VERSION : 0.7
   VAR_INPUT
      MotorStarterID : Hw_Any;   // The ID of the motor starter to read the records from
      "FB Mode" : Int;
      ManualMode : Bool;   // Used only for FB_Mode = 1 / Manual Mode Signal
      AutoMode : Bool;   // Used only for FB_Mode = 1 / Auto Mode Signal
      Interlock : Bool;   // Interlock
      AutoOn : Bool;
      HandOn : Bool;   // Hand ON
      HandOff : Bool;   // Hand OFF
      SpareIN_1 : Bool;   // Spare
      RemoteFeedbackStat : Bool;   // Status - Remote Mode Feedback
      OnStatus : Bool;   // Status - On
      DeviceOStatus : Bool;   // Status - Device Ok
      CoolindDownPeriodStatus : Bool;   // Status - Cooling Down Period Active
      EmergencyStartExecStatus : Bool;   // Status - Emergency Start Executed
      GeneralWarningStatus : Bool;   // Fault - General Warning
      GeneralFaultStatus : Bool;   // Fault - General Fault
      OverloadOperationEvent : Bool;   // Event - Overload Operation Fault (I>115%Is)
      OverloadFaultEvent : Bool;   // Event - Overload Fault
      UnbalanceFault : Bool;   // Event - Unbalance Fault
      OLandLossOfPhaseEvent : Bool;   // Event - Overload and Loss of Phase
      StalledRotorEvent : Bool;   // Event - Stalled Rotor
      HardwareFaultBasicUnitTrip : Bool;   // Trip - Hardware Fault Basic Unit
      ModuleFaultTrip : Bool;   // Trip - Module Fault
      ExecOnCommandTrip : Bool;   // Trip - Execution On-Command
      RemainingCooldDownPeriod : Int;   // Remaining Cool Down Period
      FullLoadAmps : Real;   // Full Load Amps
   END_VAR
   VAR_OUTPUT
      SpareOUT_1 : Bool;
      Stop_CMD : Bool;   // Stop Command for the Semicode
      Start_CMD : Bool;   // Start Command for the Semicode
      TestSimocode : Bool;   // Simocode Test
      EmergenyStart : Bool;   // Emergency Start
      RemoteCommandsEnabled : Bool;   // Auto Mode / Enable Remote Commands
      ResetSimocode : Bool;   // Simocode Reset
      SpareOUT_2 : Bool;
      SpareOUT_3 : Bool;
      SpareOUT_4 : Bool;
      SpareOUT_5 : Bool;
      SpareOUT_6 : Bool;
      SpareOUT_7 : Bool;
      SpareOUT_8 : Bool;
      SpareOUT_9 : Bool;
      SpareOUT_10 : Bool;
      SpareOUTW_1 : Int;
      SpareOUTW_2 : Int;
   END_VAR
   VAR
      HMI : Struct
         Controls : Struct
            Start : Bool;
            Stop : Bool;
            Reset : Bool;
            PLCMOHR : Bool;   // PLC Motor Operating Hours Reset
         END_STRUCT;
         Status : Struct
            Mode : Int;   // Simocode Mode
            MotorOperatingHours : Real;   // True Semicode Motor Operating Hours
            DeviceOperatingHours : Real;
            LMOH : Real;   // Last Motor Operating Hours
            RemainingCoolDownPeriod : Int;   // Remaining Cooldown Period
            MaxNumberOLtrips : Int;   // Maximum Number of Overload Trips
            ControlStatusWord : Word;   // Control/Status Information Bits
            MaxCurrent : Real;   // Maximum Current (Is %)
            Current1 : Real;   // Leg 1 Current (Is %)
            Current2 : Real;   // Leg 2 Current (Is %)
            Current3 : Real;   // Leg 3 Current (Is %)
            LastTripCurrent : Real;   // Last Trip Current (% of Is)
            CommandSimocode : Bool;   // Commanding Simocode to Start
         END_STRUCT;
         Config : Struct
            "RemainingCoolDownPeriod.SP" : Int := 300;
            Start_PT : Time := T#500MS;
            Stop_PT : Time := T#500MS;
         END_STRUCT;
         Math : Struct
            MOH1 : DInt;
            MOH2 : Real;
            PLCMOH : Real;   // PLC Motor Operating Hours
            LMOH : Real;
         END_STRUCT;
      END_STRUCT;
      OS : Struct
         RON : Bool;   // Remote / HMI On
         ROFF : Bool;   // Remote / HMI Off
         HON : Bool;   // Hand/Local On
         HOFF : Bool;   // Hand/Local Off
         PLCMOHR : Bool;
         LMOH1 : Bool;
         LMOH2 : Bool;
         RST : Bool;   // Reset Semicode
      END_STRUCT;
      "DS94 Record" : Struct
         "Phase Current L1 %" : USInt;
         "Phase Current L2 %" : USInt;
         "Phase Current L3 %" : USInt;
         Reserved_3 : Byte;
         "Remaining cool-down time of the motor" : UInt;
         "Motor heating_6" : USInt;
         Unbalance : USInt;
         "Motor Heating" : UInt;
         Reserved_10 : Byte;
         Reserved_11 : Byte;
         Reserved_12 : Byte;
         Reserved_13 : Byte;
         Reserved_14 : Byte;
         Reserved_15 : Byte;
         Reserved_16 : Byte;
         Reserved_17 : Byte;
         Reserved_18 : Byte;
         Reserved_19 : Byte;
         Reserved_20 : Byte;
         Reserved_21 : Byte;
         Reserved_22 : Byte;
         Reserved_23 : Byte;
         Reserved_24 : Byte;
         Reserved_25 : Byte;
         Reserved_26 : Byte;
         Reserved_27 : Byte;
         "Phase Current L1 (rms)" : UDInt;
         "Phase Current L2 (rms)" : UDInt;
         "Phase Current L3 (rms)" : UDInt;
         "Electronics Supply Voltage" : UInt;
         Reserved_42 : Byte;
         Reserved_43 : Byte;
         Reserved_44 : Byte;
         Reserved_45 : Byte;
         Reserved_46 : Byte;
         Reserved_47 : Byte;
         Reserved_48 : Byte;
         Reserved_49 : Byte;
         Reserved_50 : Byte;
         Reserved_51 : Byte;
         Reserved_52 : Byte;
         Reserved_53 : Byte;
         Reserved_54 : Byte;
         Reserved_55 : Byte;
         Reserved_56 : Byte;
         Reserved_57 : Byte;
         Reserved_58 : Byte;
         Reserved_59 : Byte;
         Reserved_60 : Byte;
         Reserved_61 : Byte;
         Reserved_62 : Byte;
         Reserved_63 : Byte;
      END_STRUCT;
      "DS94 Record_1" : Struct
         "Phase Current L1 %" : USInt;
         "Phase Current L2 %" : USInt;
         "Phase Current L3 %" : USInt;
         Reserved_3 : Byte;
         "Remaining cool-down time of the motor" : UInt;
         "Motor heating_6" : USInt;
         "Asymmetry value_7" : USInt;
         Reserved_8 : Byte;
         Reserved_9 : Byte;
         Reserved_10 : Byte;
         Reserved_11 : Byte;
         Reserved_12 : Byte;
         Reserved_13 : Byte;
         Reserved_14 : Byte;
         Reserved_15 : Byte;
         Reserved_16 : Byte;
         Reserved_17 : Byte;
         Reserved_18 : Byte;
         Reserved_19 : Byte;
         Reserved_20 : Byte;
         Reserved_21 : Byte;
         Reserved_22 : Byte;
         Reserved_23 : Byte;
         Reserved_24 : Byte;
         Reserved_25 : Byte;
         Reserved_26 : Byte;
         Reserved_27 : Byte;
         "Phase Current L1 (rms)" : UDInt;
         "Phase Current L2 (rms)" : UDInt;
         "Phase Current L3 (rms)" : UDInt;
         "Electronics Supply Voltage" : USInt;
         Reserved_46 : Byte;
         Reserved_47 : Byte;
         Reserved_48 : Byte;
         Reserved_49 : Byte;
         Reserved_50 : Byte;
         Reserved_51 : Byte;
         Reserved_52 : Byte;
         Reserved_53 : Byte;
         Reserved_54 : Byte;
         Reserved_55 : Byte;
         Reserved_56 : Byte;
         Reserved_57 : Byte;
         Reserved_58 : Byte;
         Reserved_59 : Byte;
         Reserved_60 : Byte;
         Reserved_61 : Byte;
         Reserved_62 : Byte;
      END_STRUCT;
      "DS95 Record" : Struct
         Reserved_0 : USInt;
         "Reserved_1.0" : Bool;
         "Reserved_1.1" : Bool;
         "Reserved_1.2" : Bool;
         "Reserved_1.3" : Bool;
         "Reserved_1.4" : Bool;
         "Reserved_1.5" : Bool;
         "Reserved_1.6" : Bool;
         "Reserved_1.7" : Bool;
         Reserved_2 : Byte;
         Reserved_3 : Byte;
         "Device operating hours in seconds" : UDInt;
         "Number of motor CW starts" : UDInt;
         "Number of starts motor CCW" : UDInt;
         "Number of motor overload trips" : UInt;
         Reserved_18 : Byte;
         Reserved_19 : Byte;
         "Motor current_20..23" : UDInt;
         "Last tripping current_24..27" : DInt;
         "Motor operating hours in seconds_28...31" : UDInt;
         Reserved_32 : Byte;
         Reserved_33 : Byte;
         Reserved_34 : Byte;
         Reserved_35 : Byte;
         Reserved_36 : Byte;
         Reserved_37 : Byte;
         Reserved_38 : Byte;
         Reserved_39 : Byte;
         Reserved_40 : Byte;
         Reserved_41 : Byte;
         Reserved_42 : Byte;
         Reserved_43 : Byte;
         Reserved_44 : Byte;
         Reserved_45 : Byte;
         Reserved_46 : Byte;
         Reserved_47 : Byte;
         Reserved_48 : Byte;
         Reserved_49 : Byte;
         "Number of switching element" : UInt;
         "Number of hard switching" : UInt;
         Reserved_54 : Byte;
         Reserved_55 : Byte;
         Reserved_56 : Byte;
         Reserved_57 : Byte;
         Reserved_58 : Byte;
         Reserved_59 : Byte;
         Reserved_60 : Byte;
         Reserved_61 : Byte;
         Reserved_62 : Byte;
         Reserved_63 : Byte;
         Reserved_64 : Byte;
         Reserved_65 : Byte;
         Reserved_66 : Byte;
         Reserved_67 : Byte;
         Reserved_68 : Byte;
         Reserved_69 : Byte;
         Reserved_70 : Byte;
         Reserved_71 : Byte;
         Reserved_72 : Byte;
         Reserved_73 : Byte;
         Reserved_74 : Byte;
         Reserved_75 : Byte;
         Reserved_76 : Byte;
         Reserved_77 : Byte;
         Reserved_78 : Byte;
         Reserved_79 : Byte;
         Reserved_80 : Byte;
         Reserved_81 : Byte;
         Reserved_82 : Byte;
         Reserved_83 : Byte;
         Reserved_84 : Byte;
         Reserved_85 : Byte;
         Reserved_86 : Byte;
         Reserved_87 : Byte;
         Reserved_88 : Byte;
         Reserved_89 : Byte;
      END_STRUCT;
      START_CMD_TOF : TOF_TIME;   // Start Semicode
      STOP_CMD_TOF : TOF_TIME;
      Current_RDREC : RDREC;
      Time_RDREC : RDREC;
      RDREC_REQ : SInt;
      Current_Error : SInt;
      Time_Error : SInt;
      flnk : Array[0..2] of Bool;
   END_VAR
   VAR_TEMP
      IL1_Math2 : Real;
      IL1_Math3 : Real;
      IL2_Math2 : Real;
      IL2_Math3 : Real;
      IL3_Math2 : Real;
      IL3_Math3 : Real;
      MC_Math1 : DInt;
      MC_Math2 : Real;
      MC_Math3 : Real;
      LTC_Math2 : Real;
      LTC_Math3 : Real;
      Start : Bool;
      Fault : Bool;
      "Valid Current" : Bool;
      "Valid Time" : Bool;
      MOTS : Real;   // Motor Operating Time in Seconds
      DOTH : Real;   // Device Operating Time in Hours
      DOTS : Real;   // Device Operating Time in Seconds
      MOTH : Real;   // Motor Operating Time in hours
   END_VAR
   VAR_TEMP   // added for the SCL form of the ladder/FBD networks
      _w1 : Bool;
      _w2 : Bool;
      _w3 : Bool;
      _w4 : Bool;
      _w5 : Bool;
   END_VAR
BEGIN

REGION Network 1: Read request
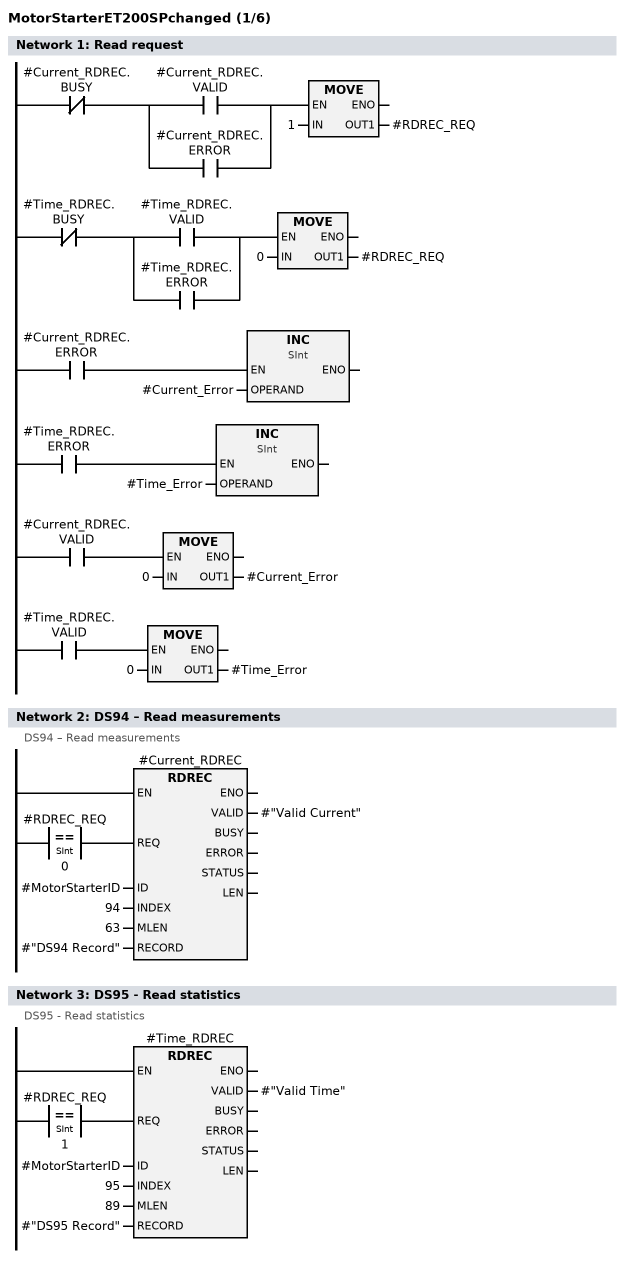
   RUNG wire#powerrail
      I_Contact( #Current_RDREC.BUSY )
      wire#w1
      Contact( #Current_RDREC.VALID )
      wire#w2
      Move(in := 1, out1 => #RDREC_REQ)
   END_RUNG
   RUNG wire#w1
      Contact( #Current_RDREC.ERROR )
   END_RUNG wire#w2
   RUNG wire#powerrail
      I_Contact( #Time_RDREC.BUSY )
      wire#w3
      Contact( #Time_RDREC.VALID )
      wire#w4
      Move(in := 0, out1 => #RDREC_REQ)
   END_RUNG
   RUNG wire#w3
      Contact( #Time_RDREC.ERROR )
   END_RUNG wire#w4
   RUNG wire#powerrail
      Contact( #Current_RDREC.ERROR )
      { S7_Templates := "DestType := SInt" } Inc( #Current_Error )
   END_RUNG
   RUNG wire#powerrail
      Contact( #Time_RDREC.ERROR )
      { S7_Templates := "DestType := SInt" } Inc( #Time_Error )
   END_RUNG
   RUNG wire#powerrail
      Contact( #Current_RDREC.VALID )
      Move(in := 0, out1 => #Current_Error)
   END_RUNG
   RUNG wire#powerrail
      Contact( #Time_RDREC.VALID )
      Move(in := 0, out1 => #Time_Error)
   END_RUNG
   // the same network as SCL:
   IF NOT #Current_RDREC.BUSY AND (#Current_RDREC.VALID OR #Current_RDREC.ERROR) THEN
       #RDREC_REQ := 1;
   END_IF;
   IF NOT #Time_RDREC.BUSY AND (#Time_RDREC.VALID OR #Time_RDREC.ERROR) THEN #RDREC_REQ := 0; END_IF;
   IF #Current_RDREC.ERROR THEN #Current_Error := #Current_Error + 1; END_IF;
   IF #Time_RDREC.ERROR THEN #Time_Error := #Time_Error + 1; END_IF;
   IF #Current_RDREC.VALID THEN #Current_Error := 0; END_IF;
   IF #Time_RDREC.VALID THEN #Time_Error := 0; END_IF;
END_REGION

REGION Network 2: DS94 – Read measurements
   // DS94 – Read measurements
   #Current_RDREC(REQ := #RDREC_REQ = 0,   // RDREC
                  ID := #MotorStarterID,
                  INDEX := 94,
                  MLEN := 63,
                  RECORD := #"DS94 Record",
                  VALID => #"Valid Current");
END_REGION

REGION Network 3: DS95 - Read statistics
   // DS95 - Read statistics
   #Time_RDREC(REQ := #RDREC_REQ = 1,   // RDREC
               ID := #MotorStarterID,
               INDEX := 95,
               MLEN := 89,
               RECORD := #"DS95 Record",
               VALID => #"Valid Time");
END_REGION

REGION Network 4: HOA in Off
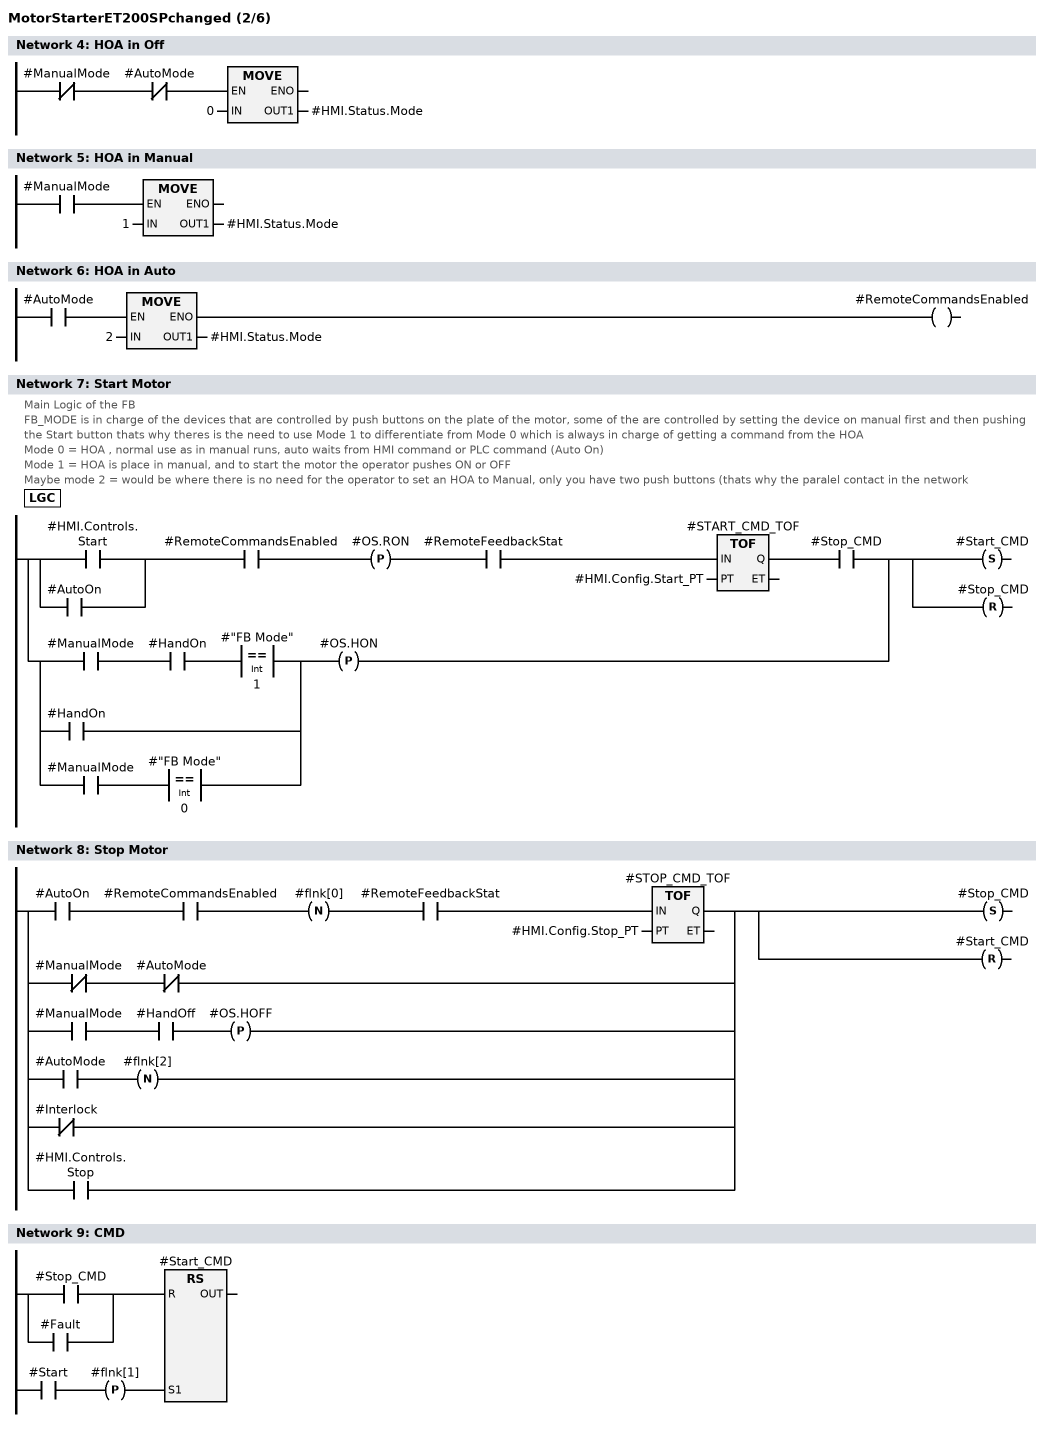
   RUNG wire#powerrail
      I_Contact( #ManualMode )
      I_Contact( #AutoMode )
      { S7_GenerateENO := "TRUE" } Move(in := 0, out1 => #HMI.Status.Mode)
   END_RUNG
   // the same network as SCL:
   IF NOT #ManualMode AND NOT #AutoMode THEN #HMI.Status.Mode := 0; END_IF;
END_REGION

REGION Network 5: HOA in Manual
   RUNG wire#powerrail
      Contact( #ManualMode )
      { S7_GenerateENO := "TRUE" } Move(in := 1, out1 => #HMI.Status.Mode)
   END_RUNG
   // the same network as SCL:
   IF #ManualMode THEN #HMI.Status.Mode := 1; END_IF;
END_REGION

REGION Network 6: HOA in Auto
   RUNG wire#powerrail
      Contact( #AutoMode )
      { S7_GenerateENO := "TRUE" } Move(in := 2, out1 => #HMI.Status.Mode)
      Coil( #RemoteCommandsEnabled )
   END_RUNG
   // the same network as SCL:
   // ENO of a box is taken as its EN; it also drops when the box reports an error
   IF #AutoMode THEN #HMI.Status.Mode := 2; END_IF;
   #RemoteCommandsEnabled := #AutoMode;
END_REGION

REGION Network 7: Start Motor
   // Main Logic of the FB
   // FB_MODE is in charge of the devices that are controlled by push buttons on the plate of the motor, some of the are controlled by setting the device on manual first and then pushing the Start button thats why theres is the need to use Mode 1 to differentiate from Mode 0 which is always in charge of getting a command from the HOA
   // Mode 0 = HOA , normal use as in manual runs, auto waits from HMI command or PLC command (Auto On)
   // Mode 1 = HOA is place in manual, and to start the motor the operator pushes ON or OFF
   // Maybe mode 2 = would be where there is no need for the operator to set an HOA to Manual, only you have two push buttons (thats why the paralel contact in the network
   LGC:
   #_w1 := (#HMI.Controls.Start OR #AutoOn) AND #RemoteCommandsEnabled;
   #_w2 := #_w1 AND NOT #OS.RON;   // rising edge
   #OS.RON := #_w1;
   #START_CMD_TOF(IN := #_w2 AND #RemoteFeedbackStat, PT := #HMI.Config.Start_PT);   // TOF
   #_w3 := (#ManualMode AND #HandOn AND (#"FB Mode" = 1)) OR #HandOn OR (#ManualMode AND (#"FB Mode" = 0));
   #_w4 := #_w3 AND NOT #OS.HON;   // rising edge
   #OS.HON := #_w3;
   IF (#START_CMD_TOF.Q AND #Stop_CMD) OR #_w4 THEN
       #Start_CMD := TRUE;
       #Stop_CMD := FALSE;
   END_IF;
END_REGION

REGION Network 8: Stop Motor
   #_w1 := #AutoOn AND #RemoteCommandsEnabled;
   #_w2 := NOT #_w1 AND #flnk[0];   // falling edge
   #flnk[0] := #_w1;
   #STOP_CMD_TOF(IN := #_w2 AND #RemoteFeedbackStat, PT := #HMI.Config.Stop_PT);   // TOF
   #_w3 := #ManualMode AND #HandOff;
   #_w4 := #_w3 AND NOT #OS.HOFF;   // rising edge
   #OS.HOFF := #_w3;
   #_w5 := NOT #AutoMode AND #flnk[2];   // falling edge
   #flnk[2] := #AutoMode;
   IF #STOP_CMD_TOF.Q OR (NOT #ManualMode AND NOT #AutoMode) OR #_w4 OR #_w5 OR NOT #Interlock OR #HMI.Controls.Stop THEN
       #Stop_CMD := TRUE;
       #Start_CMD := FALSE;
   END_IF;
END_REGION

REGION Network 9: CMD
   RUNG wire#powerrail
      Contact( #Stop_CMD )
      wire#w1
      S_RS(operand := #Start_CMD, s1 := wire#w2)
   END_RUNG
   RUNG wire#powerrail
      Contact( #Fault )
   END_RUNG wire#w1
   RUNG wire#powerrail
      Contact( #Start )
      P_Trig( #flnk[1] )
   END_RUNG wire#w2
   // the same network as SCL:
   #_w1 := #Start AND NOT #flnk[1];   // rising edge
   #flnk[1] := #Start;
   IF #Stop_CMD OR #Fault THEN
       #Start_CMD := FALSE;   // RS flip-flop
   END_IF;
   IF #_w1 THEN #Start_CMD := TRUE; END_IF;
END_REGION

REGION Network 10: Interlock
   // Main Logic of the FB
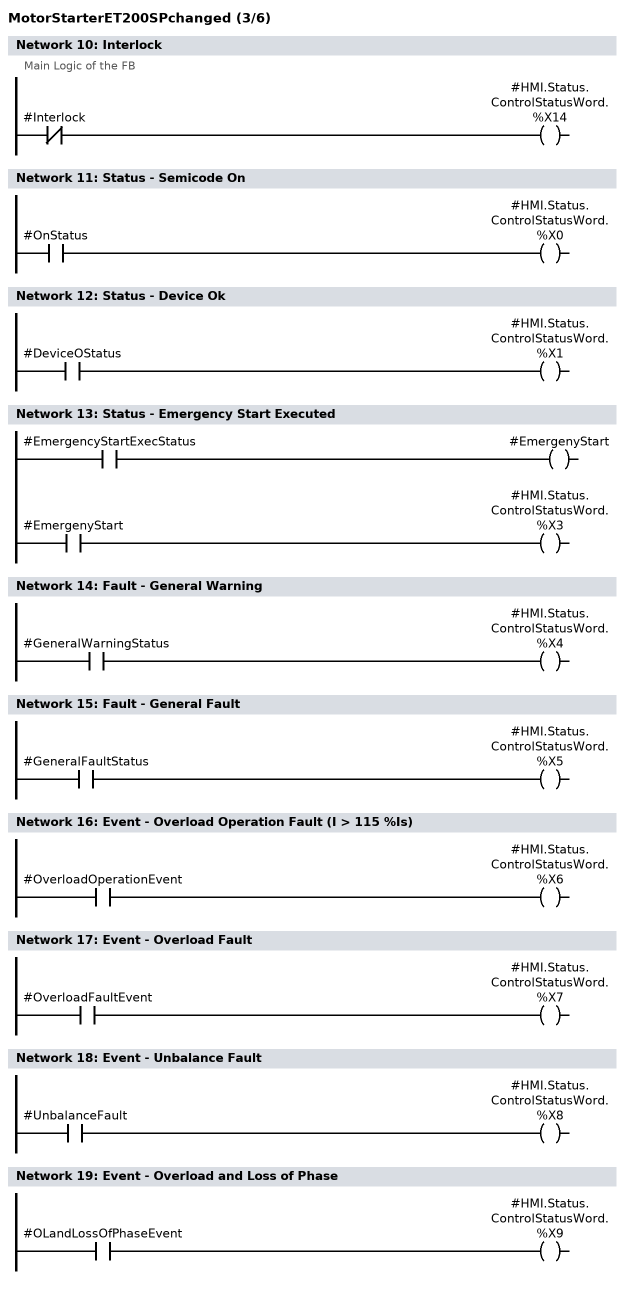
   RUNG wire#powerrail
      I_Contact( #Interlock )
      Coil( #HMI.Status.ControlStatusWord.%X14 )
   END_RUNG
   // the same network as SCL:
   #HMI.Status.ControlStatusWord.%X14 := NOT #Interlock;
END_REGION

REGION Network 11: Status - Semicode On
   RUNG wire#powerrail
      Contact( #OnStatus )
      Coil( #HMI.Status.ControlStatusWord.%X0 )
   END_RUNG
   // the same network as SCL:
   #HMI.Status.ControlStatusWord.%X0 := #OnStatus;
END_REGION

REGION Network 12: Status - Device Ok
   RUNG wire#powerrail
      Contact( #DeviceOStatus )
      Coil( #HMI.Status.ControlStatusWord.%X1 )
   END_RUNG
   // the same network as SCL:
   #HMI.Status.ControlStatusWord.%X1 := #DeviceOStatus;
END_REGION

REGION Network 13: Status - Emergency Start Executed
   RUNG wire#powerrail
      Contact( #EmergencyStartExecStatus )
      Coil( #EmergenyStart )
   END_RUNG
   RUNG wire#powerrail
      Contact( #EmergenyStart )
      Coil( #HMI.Status.ControlStatusWord.%X3 )
   END_RUNG
   // the same network as SCL:
   #EmergenyStart := #EmergencyStartExecStatus;
   #HMI.Status.ControlStatusWord.%X3 := #EmergenyStart;
END_REGION

REGION Network 14: Fault - General Warning
   RUNG wire#powerrail
      Contact( #GeneralWarningStatus )
      Coil( #HMI.Status.ControlStatusWord.%X4 )
   END_RUNG
   // the same network as SCL:
   #HMI.Status.ControlStatusWord.%X4 := #GeneralWarningStatus;
END_REGION

REGION Network 15: Fault - General Fault
   RUNG wire#powerrail
      Contact( #GeneralFaultStatus )
      Coil( #HMI.Status.ControlStatusWord.%X5 )
   END_RUNG
   // the same network as SCL:
   #HMI.Status.ControlStatusWord.%X5 := #GeneralFaultStatus;
END_REGION

REGION Network 16: Event - Overload Operation Fault (I > 115 %Is)
   RUNG wire#powerrail
      Contact( #OverloadOperationEvent )
      Coil( #HMI.Status.ControlStatusWord.%X6 )
   END_RUNG
   // the same network as SCL:
   #HMI.Status.ControlStatusWord.%X6 := #OverloadOperationEvent;
END_REGION

REGION Network 17: Event - Overload Fault
   RUNG wire#powerrail
      Contact( #OverloadFaultEvent )
      Coil( #HMI.Status.ControlStatusWord.%X7 )
   END_RUNG
   // the same network as SCL:
   #HMI.Status.ControlStatusWord.%X7 := #OverloadFaultEvent;
END_REGION

REGION Network 18: Event - Unbalance Fault
   RUNG wire#powerrail
      Contact( #UnbalanceFault )
      Coil( #HMI.Status.ControlStatusWord.%X8 )
   END_RUNG
   // the same network as SCL:
   #HMI.Status.ControlStatusWord.%X8 := #UnbalanceFault;
END_REGION

REGION Network 19: Event - Overload and Loss of Phase
   RUNG wire#powerrail
      Contact( #OLandLossOfPhaseEvent )
      Coil( #HMI.Status.ControlStatusWord.%X9 )
   END_RUNG
   // the same network as SCL:
   #HMI.Status.ControlStatusWord.%X9 := #OLandLossOfPhaseEvent;
END_REGION

REGION Network 20: Event - Stalled Rotor
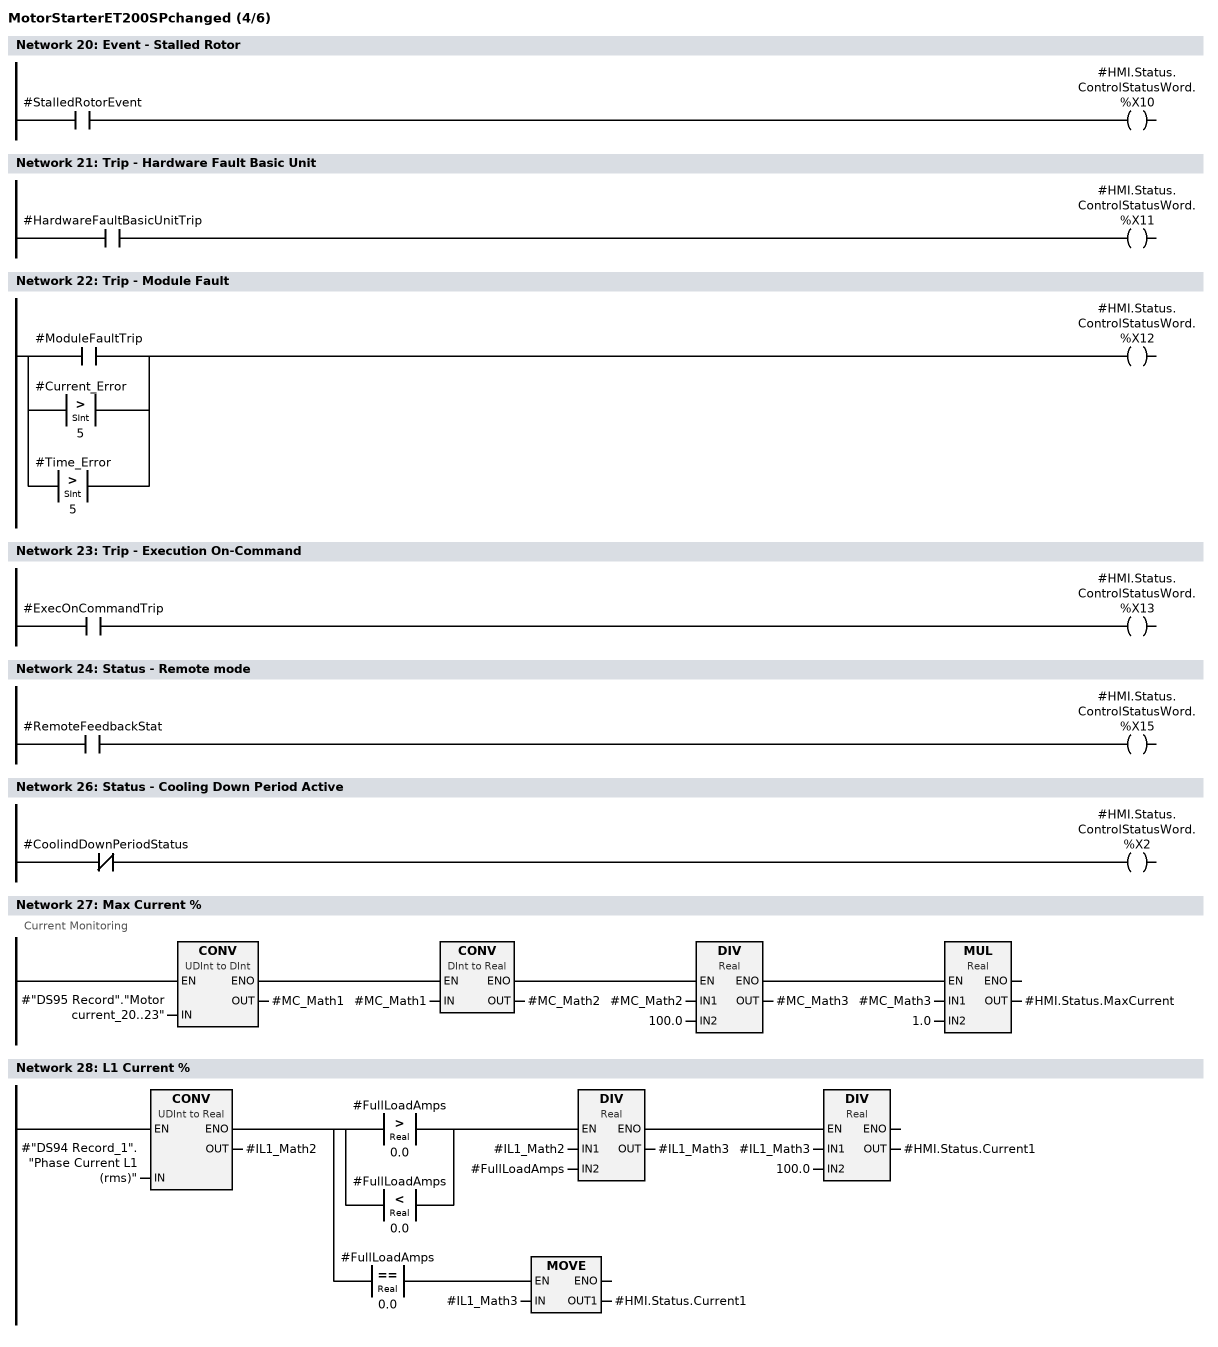
   RUNG wire#powerrail
      Contact( #StalledRotorEvent )
      Coil( #HMI.Status.ControlStatusWord.%X10 )
   END_RUNG
   // the same network as SCL:
   #HMI.Status.ControlStatusWord.%X10 := #StalledRotorEvent;
END_REGION

REGION Network 21: Trip - Hardware Fault Basic Unit
   RUNG wire#powerrail
      Contact( #HardwareFaultBasicUnitTrip )
      Coil( #HMI.Status.ControlStatusWord.%X11 )
   END_RUNG
   // the same network as SCL:
   #HMI.Status.ControlStatusWord.%X11 := #HardwareFaultBasicUnitTrip;
END_REGION

REGION Network 22: Trip - Module Fault
   RUNG wire#powerrail
      Contact( #ModuleFaultTrip )
      wire#w1
      Coil( #HMI.Status.ControlStatusWord.%X12 )
   END_RUNG
   RUNG wire#powerrail
      { S7_Templates := "SrcType := SInt" } GT_Contact(in1 := #Current_Error, in2 := 5)
   END_RUNG wire#w1
   RUNG wire#powerrail
      { S7_Templates := "SrcType := SInt" } GT_Contact(in1 := #Time_Error, in2 := 5)
   END_RUNG wire#w1
   // the same network as SCL:
   #HMI.Status.ControlStatusWord.%X12 := #ModuleFaultTrip OR (#Current_Error > 5) OR (#Time_Error > 5);
END_REGION

REGION Network 23: Trip - Execution On-Command
   RUNG wire#powerrail
      Contact( #ExecOnCommandTrip )
      Coil( #HMI.Status.ControlStatusWord.%X13 )
   END_RUNG
   // the same network as SCL:
   #HMI.Status.ControlStatusWord.%X13 := #ExecOnCommandTrip;
END_REGION

REGION Network 24: Status - Remote mode
   RUNG wire#powerrail
      Contact( #RemoteFeedbackStat )
      Coil( #HMI.Status.ControlStatusWord.%X15 )
   END_RUNG
   // the same network as SCL:
   #HMI.Status.ControlStatusWord.%X15 := #RemoteFeedbackStat;
END_REGION

REGION Network 25 (SCL): Motor Operating Hours
   #DOTS := UDINT_TO_REAL(#"DS95 Record"."Device operating hours in seconds");
   #DOTH := #DOTS / Real#3610.68;
   #MOTS := UDINT_TO_REAL(#"DS95 Record"."Motor operating hours in seconds_28...31");
   #MOTH := #MOTS / Real#6027.66;
   #HMI.Status.DeviceOperatingHours := #DOTH;
   #HMI.Status.MotorOperatingHours := #MOTH;
END_REGION

REGION Network 26: Status - Cooling Down Period Active
   RUNG wire#powerrail
      I_Contact( #CoolindDownPeriodStatus )
      Coil( #HMI.Status.ControlStatusWord.%X2 )
   END_RUNG
   // the same network as SCL:
   #HMI.Status.ControlStatusWord.%X2 := NOT #CoolindDownPeriodStatus;
END_REGION

REGION Network 27: Max Current %
   // Current Monitoring
   RUNG wire#powerrail
      { S7_Templates := "[SrcType := UDInt, DestType := DInt]"; S7_GenerateENO := "TRUE" } Convert(in := #"DS95 Record"."Motor current_20..23", out => #MC_Math1)
      { S7_Templates := "[SrcType := DInt, DestType := Real]"; S7_GenerateENO := "TRUE" } Convert(in := #MC_Math1, out => #MC_Math2)
      { S7_Templates := "SrcType := Real"; S7_GenerateENO := "TRUE" } Div(in1 := #MC_Math2, in2 := 100.0, out => #MC_Math3)
      { S7_Templates := "SrcType := Real"; S7_GenerateENO := "TRUE" } Mul(in1 := #MC_Math3, in2 := 1.0, out => #HMI.Status.MaxCurrent)
   END_RUNG
   // the same network as SCL:
   // ENO of a box is taken as its EN; it also drops when the box reports an error
   #MC_Math1 := UDINT_TO_DINT(#"DS95 Record"."Motor current_20..23");
   #MC_Math2 := DINT_TO_REAL(#MC_Math1);
   #MC_Math3 := #MC_Math2 / 100.0;
   #HMI.Status.MaxCurrent := #MC_Math3 * 1.0;
END_REGION

REGION Network 28: L1 Current %
   RUNG wire#powerrail
      { S7_Templates := "[SrcType := UDInt, DestType := Real]"; S7_GenerateENO := "TRUE" } Convert(in := #"DS94 Record_1"."Phase Current L1 (rms)", out => #IL1_Math2)
      wire#w1
      { S7_Templates := "SrcType := Real" } GT_Contact(in1 := #FullLoadAmps, in2 := 0.0)
      wire#w2
      { S7_Templates := "SrcType := Real"; S7_GenerateENO := "TRUE" } Div(in1 := #IL1_Math2, in2 := #FullLoadAmps, out => #IL1_Math3)
      { S7_Templates := "SrcType := Real"; S7_GenerateENO := "TRUE" } Div(in1 := #IL1_Math3, in2 := 100.0, out => #HMI.Status.Current1)
   END_RUNG
   RUNG wire#w1
      { S7_Templates := "SrcType := Real" } LT_Contact(in1 := #FullLoadAmps, in2 := 0.0)
   END_RUNG wire#w2
   RUNG wire#w1
      { S7_Templates := "SrcType := Real" } EQ_Contact(in1 := #FullLoadAmps, in2 := 0.0)
      Move(in := #IL1_Math3, out1 => #HMI.Status.Current1)
   END_RUNG
   // the same network as SCL:
   // ENO of a box is taken as its EN; it also drops when the box reports an error
   #IL1_Math2 := UDINT_TO_REAL(#"DS94 Record_1"."Phase Current L1 (rms)");
   IF (#FullLoadAmps > 0.0) OR (#FullLoadAmps < 0.0) THEN
       #IL1_Math3 := #IL1_Math2 / #FullLoadAmps;
       #HMI.Status.Current1 := #IL1_Math3 / 100.0;
   END_IF;
   IF #FullLoadAmps = 0.0 THEN #HMI.Status.Current1 := #IL1_Math3; END_IF;
END_REGION

REGION Network 29: L2 Current %
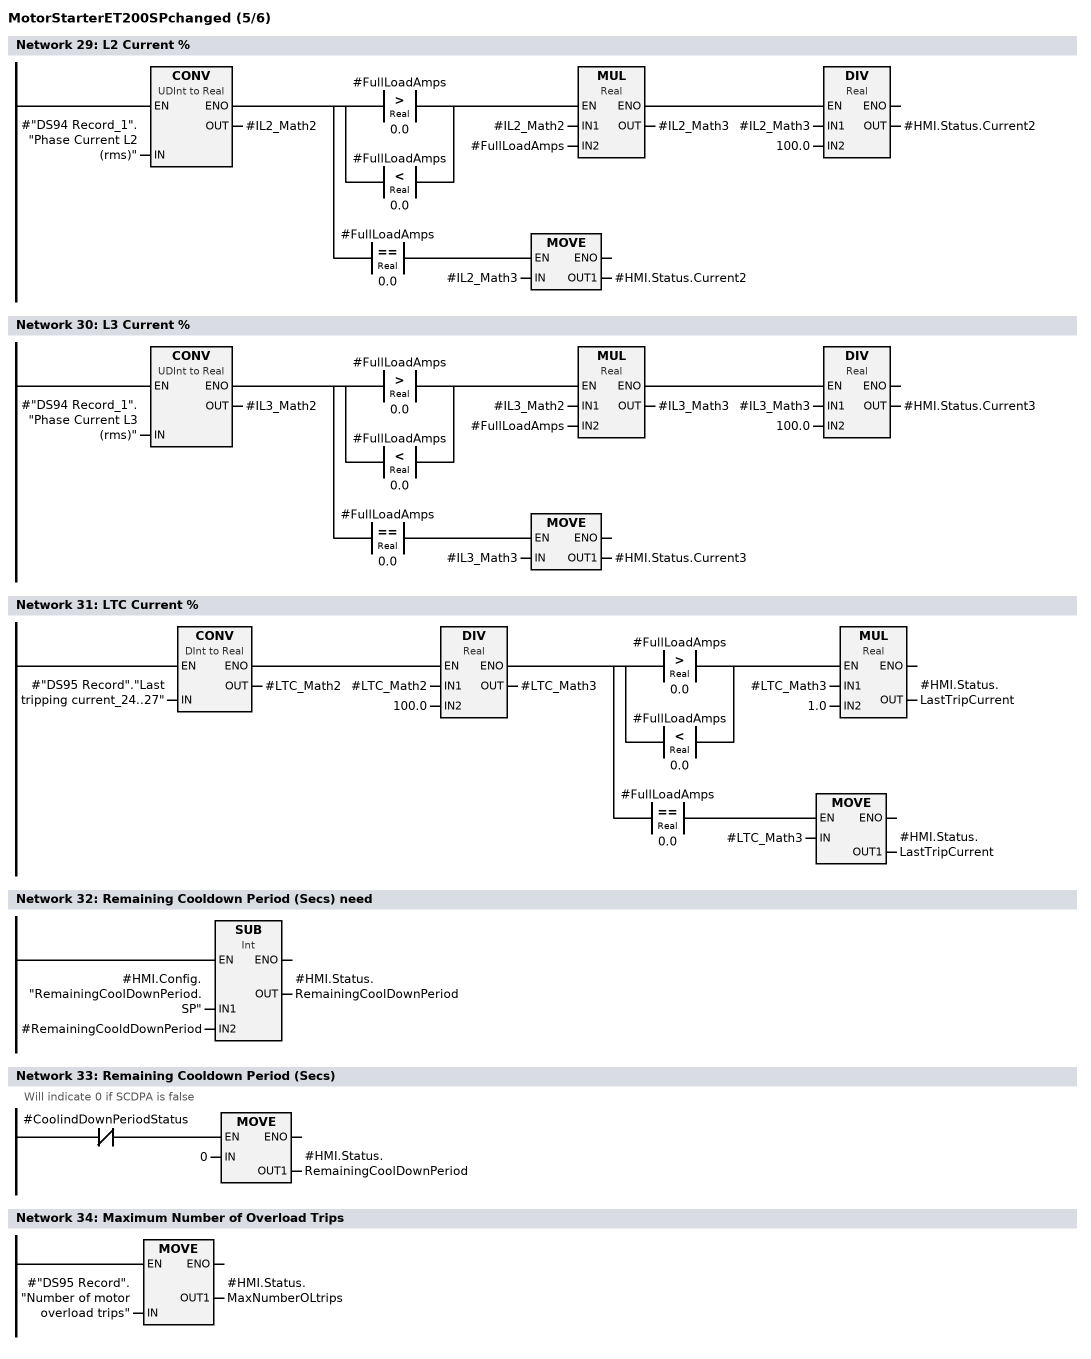
   RUNG wire#powerrail
      { S7_Templates := "[SrcType := UDInt, DestType := Real]"; S7_GenerateENO := "TRUE" } Convert(in := #"DS94 Record_1"."Phase Current L2 (rms)", out => #IL2_Math2)
      wire#w1
      { S7_Templates := "SrcType := Real" } GT_Contact(in1 := #FullLoadAmps, in2 := 0.0)
      wire#w2
      { S7_Templates := "SrcType := Real"; S7_GenerateENO := "TRUE" } Mul(in1 := #IL2_Math2, in2 := #FullLoadAmps, out => #IL2_Math3)
      { S7_Templates := "SrcType := Real"; S7_GenerateENO := "TRUE" } Div(in1 := #IL2_Math3, in2 := 100.0, out => #HMI.Status.Current2)
   END_RUNG
   RUNG wire#w1
      { S7_Templates := "SrcType := Real" } LT_Contact(in1 := #FullLoadAmps, in2 := 0.0)
   END_RUNG wire#w2
   RUNG wire#w1
      { S7_Templates := "SrcType := Real" } EQ_Contact(in1 := #FullLoadAmps, in2 := 0.0)
      Move(in := #IL2_Math3, out1 => #HMI.Status.Current2)
   END_RUNG
   // the same network as SCL:
   // ENO of a box is taken as its EN; it also drops when the box reports an error
   #IL2_Math2 := UDINT_TO_REAL(#"DS94 Record_1"."Phase Current L2 (rms)");
   IF (#FullLoadAmps > 0.0) OR (#FullLoadAmps < 0.0) THEN
       #IL2_Math3 := #IL2_Math2 * #FullLoadAmps;
       #HMI.Status.Current2 := #IL2_Math3 / 100.0;
   END_IF;
   IF #FullLoadAmps = 0.0 THEN #HMI.Status.Current2 := #IL2_Math3; END_IF;
END_REGION

REGION Network 30: L3 Current %
   RUNG wire#powerrail
      { S7_Templates := "[SrcType := UDInt, DestType := Real]"; S7_GenerateENO := "TRUE" } Convert(in := #"DS94 Record_1"."Phase Current L3 (rms)", out => #IL3_Math2)
      wire#w1
      { S7_Templates := "SrcType := Real" } GT_Contact(in1 := #FullLoadAmps, in2 := 0.0)
      wire#w2
      { S7_Templates := "SrcType := Real"; S7_GenerateENO := "TRUE" } Mul(in1 := #IL3_Math2, in2 := #FullLoadAmps, out => #IL3_Math3)
      { S7_Templates := "SrcType := Real"; S7_GenerateENO := "TRUE" } Div(in1 := #IL3_Math3, in2 := 100.0, out => #HMI.Status.Current3)
   END_RUNG
   RUNG wire#w1
      { S7_Templates := "SrcType := Real" } LT_Contact(in1 := #FullLoadAmps, in2 := 0.0)
   END_RUNG wire#w2
   RUNG wire#w1
      { S7_Templates := "SrcType := Real" } EQ_Contact(in1 := #FullLoadAmps, in2 := 0.0)
      Move(in := #IL3_Math3, out1 => #HMI.Status.Current3)
   END_RUNG
   // the same network as SCL:
   // ENO of a box is taken as its EN; it also drops when the box reports an error
   #IL3_Math2 := UDINT_TO_REAL(#"DS94 Record_1"."Phase Current L3 (rms)");
   IF (#FullLoadAmps > 0.0) OR (#FullLoadAmps < 0.0) THEN
       #IL3_Math3 := #IL3_Math2 * #FullLoadAmps;
       #HMI.Status.Current3 := #IL3_Math3 / 100.0;
   END_IF;
   IF #FullLoadAmps = 0.0 THEN #HMI.Status.Current3 := #IL3_Math3; END_IF;
END_REGION

REGION Network 31: LTC Current %
   RUNG wire#powerrail
      { S7_Templates := "[SrcType := DInt, DestType := Real]"; S7_GenerateENO := "TRUE" } Convert(in := #"DS95 Record"."Last tripping current_24..27", out => #LTC_Math2)
      { S7_Templates := "SrcType := Real"; S7_GenerateENO := "TRUE" } Div(in1 := #LTC_Math2, in2 := 100.0, out => #LTC_Math3)
      wire#w1
      { S7_Templates := "SrcType := Real" } GT_Contact(in1 := #FullLoadAmps, in2 := 0.0)
      wire#w2
      { S7_Templates := "SrcType := Real"; S7_GenerateENO := "TRUE" } Mul(in1 := #LTC_Math3, in2 := 1.0, out => #HMI.Status.LastTripCurrent)
   END_RUNG
   RUNG wire#w1
      { S7_Templates := "SrcType := Real" } LT_Contact(in1 := #FullLoadAmps, in2 := 0.0)
   END_RUNG wire#w2
   RUNG wire#w1
      { S7_Templates := "SrcType := Real" } EQ_Contact(in1 := #FullLoadAmps, in2 := 0.0)
      Move(in := #LTC_Math3, out1 => #HMI.Status.LastTripCurrent)
   END_RUNG
   // the same network as SCL:
   // ENO of a box is taken as its EN; it also drops when the box reports an error
   #LTC_Math2 := DINT_TO_REAL(#"DS95 Record"."Last tripping current_24..27");
   #LTC_Math3 := #LTC_Math2 / 100.0;
   IF (#FullLoadAmps > 0.0) OR (#FullLoadAmps < 0.0) THEN
       #HMI.Status.LastTripCurrent := #LTC_Math3 * 1.0;
   END_IF;
   IF #FullLoadAmps = 0.0 THEN #HMI.Status.LastTripCurrent := #LTC_Math3; END_IF;
END_REGION

REGION Network 32: Remaining Cooldown Period (Secs) need
   RUNG wire#powerrail
      { S7_Templates := "SrcType := Int"; S7_GenerateENO := "TRUE" } Sub(in1 := #HMI.Config."RemainingCoolDownPeriod.SP", in2 := #RemainingCooldDownPeriod, out => #HMI.Status.RemainingCoolDownPeriod)
   END_RUNG
   // the same network as SCL:
   #HMI.Status.RemainingCoolDownPeriod := #HMI.Config."RemainingCoolDownPeriod.SP" - #RemainingCooldDownPeriod;
END_REGION

REGION Network 33: Remaining Cooldown Period (Secs)
   // Will indicate 0 if SCDPA is false
   RUNG wire#powerrail
      I_Contact( #CoolindDownPeriodStatus )
      { S7_GenerateENO := "TRUE" } Move(in := 0, out1 => #HMI.Status.RemainingCoolDownPeriod)
   END_RUNG
   // the same network as SCL:
   IF NOT #CoolindDownPeriodStatus THEN #HMI.Status.RemainingCoolDownPeriod := 0; END_IF;
END_REGION

REGION Network 34: Maximum Number of Overload Trips
   RUNG wire#powerrail
      { S7_GenerateENO := "TRUE" } Move(in := #"DS95 Record"."Number of motor overload trips", out1 => #HMI.Status.MaxNumberOLtrips)
   END_RUNG
   // the same network as SCL:
   #HMI.Status.MaxNumberOLtrips := #"DS95 Record"."Number of motor overload trips";
END_REGION

REGION Network 35: Simocode Reset Commands
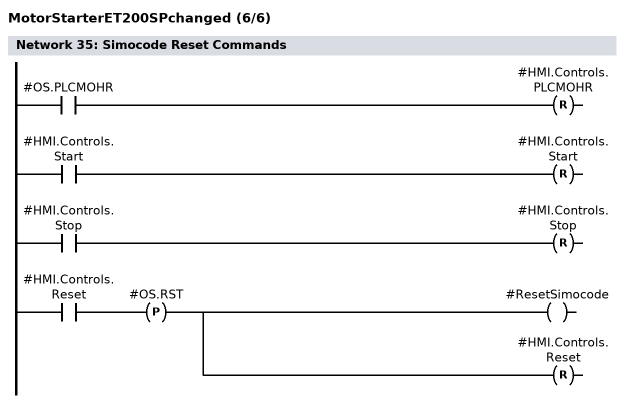
   RUNG wire#powerrail
      Contact( #OS.PLCMOHR )
      R_Coil( #HMI.Controls.PLCMOHR )
   END_RUNG
   RUNG wire#powerrail
      Contact( #HMI.Controls.Start )
      R_Coil( #HMI.Controls.Start )
   END_RUNG
   RUNG wire#powerrail
      Contact( #HMI.Controls.Stop )
      R_Coil( #HMI.Controls.Stop )
   END_RUNG
   RUNG wire#powerrail
      Contact( #HMI.Controls.Reset )
      P_Trig( #OS.RST )
      wire#w1
      Coil( #ResetSimocode )
   END_RUNG
   RUNG wire#w1
      R_Coil( #HMI.Controls.Reset )
   END_RUNG
   // the same network as SCL:
   IF #OS.PLCMOHR THEN #HMI.Controls.PLCMOHR := FALSE; END_IF;
   IF #HMI.Controls.Start THEN #HMI.Controls.Start := FALSE; END_IF;
   IF #HMI.Controls.Stop THEN #HMI.Controls.Stop := FALSE; END_IF;
   #_w1 := #HMI.Controls.Reset AND NOT #OS.RST;   // rising edge
   #OS.RST := #HMI.Controls.Reset;
   #ResetSimocode := #_w1;
   IF #_w1 THEN #HMI.Controls.Reset := FALSE; END_IF;
END_REGION
END_FUNCTION_BLOCK

// folder: 1}Library/PID

FUNCTION_BLOCK "PID_SSAC"   // FB1, LAD
{ S7_Optimized_Access := 'TRUE' }
VERSION : 0.1
   VAR_INPUT
      processVariable : Real;
      processVariableLowerLimit : Real;
      processVariableUpperLimit : Real;
      notInhibited : Bool := TRUE;
      remoteSetpoint : Real;
      enableManualMode : Bool;
      enableRemoteSetpoint : Bool;
   END_VAR
   VAR_OUTPUT
      scaledInput : Real;
      output : Real;   // Manipulated Value REAL
      outputPer : Int;   // Manipulated Value INT
      outputPwm : Bool;   // Output PWM
   END_VAR
   VAR_IN_OUT
      pid : PID_Compact;
   END_VAR
   VAR RETAIN
      hmi : Struct
         Controls : Struct
            setpoint : Real;   // Setpoint sent to PID
            manualEnable : Bool;   // Enables Manual mode
            manualOutput : Real;   // Manual Output sent to PID 0 to 100 %
            remoteEnable : Bool;
            resetController : Bool;   // Resets Controller sent to PID
            resetError : Bool;   // ErrorAck to PID
            modeActivate : Bool;   // Execute the change of mode
         END_STRUCT;
         Config : Struct
            P : Real := 0.1;   // Proportional Control sent to PID
            I : Real := 10.0;   // Integral Control sent to PID
            D : Real := 0.0;   // Derivative Control sent to PID
            OutputHighLimit : Real := 100.0;   // Output Upper Limit sent to PID
            OutputLowLimit : Real := 0.0;   // Output Lower Limit sent to PID
            rampDownTime : Real := 1.0;
            rampUpTime : Real := 1.0;
            allowPvFaultOverride : Bool;   // Allows operator to override PV fault
            rampSetpointEnabled : Bool;   // Enables the ramping of a setpoint inside the PID
            rampSetpointValue : Real;   // Value to be reached in the ramp
            inhibitedOutput : Real := 0.0;   // Inhibited Value set by the Operator 0 to 100
            mode : Int := 4;   // Mode selected by operator 1=pretune,2=finetuning,3=automatic,4-manual, 5-Substitute output, 6-Remote
            deviationSetpoint : Real := 100.0;   // Deviation of Setpoint vs PV
         END_STRUCT;
         Status : Struct
            output : Real;
            processVariable : Real;
            faulted : Bool;   // Transmitter Faulted
            notInhibited : Bool;   // PID inhibited (interlocked, off)
            pidState : Int;   // Current mode of operation (0-Inactive, 1-SUT, 2-TIR, 3-Automatic, 4-Manual, 5-Substitute output)
         END_STRUCT;
         Alarms : Struct
            errorWord : DWord;   // Error Word of PID
            error : Bool;   // Error in PID
            deviation : Bool;   // Deviation Alarm true when deviated
         END_STRUCT;
      END_STRUCT;
   END_VAR
   VAR
      triggers : Array[0..20] of Bool;
      instanceSetpointRamp : RampFunction;
      inputManunalFlag : Bool;
      inputRemoteFlag : Bool;
      "Split Range 'V'" : "Split Range 'V'";
      deviatonAlarmDelay : TON_TIME;
   END_VAR
   VAR_TEMP
      tempDeviationAbs : Real;
   END_VAR
   VAR_TEMP   // added for the SCL form of the ladder/FBD networks
      _w1 : Bool;
      _w2 : Bool;
      _w3 : Bool;
      _w4 : Bool;
      _w5 : Bool;
   END_VAR
BEGIN

REGION Network 1: Mode of PID
   // Current mode of operation (0-Inactive, 1-PreTunning, 2-FineTunning, 3-Automatic, 4-Manual, 5-Substitute output)